// TIA Portal project "Lagerregal_3" (V20)

(* hardware
DEVICE "S7-1500/ET200MP-Station_1"  S7-1500 station
   slot 0: "Profilschiene_0"  Rack  6ES7 590-1***0-0AA0
   slot 1: "PLC_1"  CPU 1513-1 PN  6ES7 513-1AM03-0AB0  V4.0
      slot 3: "CPU-Display_1"  6ES7591-1AA00-0AA0
      slot 32768: "PROFINET-Schnittstelle_1"  X1
         slot 32769: "Port_1"  X1 P1
         slot 32770: "Port_2"  X1 P2
      slot 34817: "Virtual CP interface port_1"  Virtual CP interface port  Virtual CP interface port FW V4.0
   slot 2: "DI 16x24VDC BA_1"  DI 16x24VDC BA  6ES7 521-1BH10-0AA0  V1.1
   slot 3: "DQ 16x24VDC/0.5A ST_1"  DQ 16x24VDC/0.5A ST  6ES7 522-1BH00-0AB0  V2.0
   slot 4: "AI 8xU/I/R/RTD BA_2"  AI 8xU/I/R/RTD BA  6ES7 531-7QF00-0AB0  V1.0
   slot 5: "AI 8xU/I/R/RTD BA_1"  AI 8xU/I/R/RTD BA  6ES7 531-7QF00-0AB0  V1.0
DEVICE "HMI_1"  TP700 Comfort
   slot 0: "HMI_1"  TP700 Comfort  6AV2 124-0GC01-0AX0  17.0.0.0
   slot 1: "HMI_RT_1"  TP700 Comfort  6AV2 124-0GC01-0AX0  17.0.0.0
   slot 5: "HMI_1.IE_CP_1"  PROFINET Interface  17.0.0.0
      slot 1: "PROFINET Schnittstelle_1"  PROFINET Interface
         slot 1: "Port_1"  Port
         slot 2: "Port_2"  Port
   slot 7: "HMI_1.MPI/DP_CP_1"  MPI/DP Interface  17.0.0.0
*)

// ===== PLC "PLC_1"  CPU 1513-1 PN =====

VAR_GLOBAL   // PLC tag table "Standard-Variablentabelle"
   "Clock_Byte" AT %MB0 : Byte;
   "Clock_10Hz" AT %M0.0 : Bool;
   "Clock_5Hz" AT %M0.1 : Bool;
   "Clock_2.5Hz" AT %M0.2 : Bool;
   "Clock_2Hz" AT %M0.3 : Bool;
   "Clock_1.25Hz" AT %M0.4 : Bool;
   "Clock_1Hz" AT %M0.5 : Bool;
   "Clock_0.625Hz" AT %M0.6 : Bool;
   "Clock_0.5Hz" AT %M0.7 : Bool;
END_VAR

VAR_GLOBAL CONSTANT   // PLC tag table "Standard-Variablentabelle"
   "Fachhoehe" : Int := 4800;
   "Fachbreite" : Int := 2962;
   "Offset-Z" : Int := 1800;
   "Offset-X" : Int := 3952;
   "Faecher_pro_Zeile" : Int := 9;
   "Faecher_pro_Spalte" : Int := 6;
   "Anheben_Absenken" : Int := 1000;
END_VAR

VAR_GLOBAL   // PLC tag table "Eingaenge"
   "S1" AT %I0.0 : Bool;   // Not-Aus
   "S2" AT %I0.1 : Bool;   // Anlage ein
   "S3" AT %I0.2 : Bool;   // Starttaster
   "1B1" AT %I0.3 : Bool;   // Sensor 1. Einlassband Anfang
   "1B2" AT %I0.4 : Bool;   // Sensor 1. Einlassband Ende
   "2B1" AT %I0.5 : Bool;   // Sensor 2. Einlassband Anfang
   "2B2" AT %I0.6 : Bool;   // Sensor 2. Einlassband Ende
   "3B1" AT %I0.7 : Bool;   // Sensor 3. Einlassband
   "4B1" AT %I1.0 : Bool;   // Sensor 1. Auslassband
   "5B1" AT %I1.1 : Bool;   // Sensor 2. Auslassband
   "6B1" AT %I1.2 : Bool;   // Endlage Gabel-Kran 1 (links)
   "6B2" AT %I1.3 : Bool;   // Endlage Gabel-Kran 1 (rechts)
   "6B3" AT %I1.4 : Bool;   // Endlage Gabel-Kran 1 (mitte)
   "7B1" AT %I1.5 : Bool;   // Endlage Gabel-Kran 2 (links)
   "7B2" AT %I1.6 : Bool;   // Endlage Gabel-Kran 2 (rechts)
   "7B3" AT %I1.7 : Bool;   // Endlage Gabel-Kran 2 (mitte)
   "2B3" AT %EW30 : Int;   // Kamera am Einlass (Bauteilerkennung)
   "6B4" AT %EW32 : Int;   // X-Achse Kran 1 Ist-Pos
   "6B5" AT %EW34 : Int;   // Z-Achse Kran 1 Ist-Pos
   "7B4" AT %EW36 : Int;   // X-Achse Kran 2 Ist-Pos
   "7B5" AT %EW38 : Int;   // Z-Achse Kran 2 Ist-Pos
END_VAR

VAR_GLOBAL   // PLC tag table "Ausgaenge"
   "H3" AT %Q0.2 : Bool;   // Starttasterleuchte
   "1M1" AT %Q0.3 : Bool;   // 1. Einlassband
   "2M1" AT %Q0.5 : Bool;   // 2. Einlassband
   "3M1" AT %Q0.7 : Bool;   // 3. Einlassband
   "4M1" AT %Q1.0 : Bool;   // 1. Auslassband
   "5M1" AT %Q1.1 : Bool;   // 2. Auslassband
   "6M1" AT %Q1.2 : Bool;   // Gabel-Kran 1 (links)
   "6M2" AT %Q1.3 : Bool;   // Gabel-Kran 1 (rechts)
   "7M1" AT %Q1.5 : Bool;   // Gabel-Kran 2 (links)
   "7M2" AT %Q1.6 : Bool;   // Gabel-Kran 2 (rechts)
   "6M4" AT %AW32 : Int;   // X-Achse Kran 1 Soll-Pos
   "6M5" AT %AW34 : Int;   // Z-Achse Kran 1 Soll-Pos
   "7M4" AT %AW36 : Int;   // X-Achse Kran 2 Soll-Pos
   "7M5" AT %AW38 : Int;   // Z-Achse Kran 2 Soll-Pos
END_VAR

TYPE "typKran_Pos"
   STRUCT
      "X-Ist" : Int;
      "X-Soll" : Int;
      "Z-Ist" : Int;
      "Z-Soll" : Int;
   END_STRUCT;
END_TYPE

TYPE "typLagerplatz"
   STRUCT
      Flags : Struct
         Belegt : Bool;
         In_Benutzung : Bool;
      END_STRUCT;
   END_STRUCT;
END_TYPE

TYPE "typSchritte"
   STRUCT
      Schritt_Init : Bool;
      Kran : Struct
         Schritt_1 : Bool;
         Schritt_2 : Bool;
         Schritt_3 : Bool;
         Schritt_4 : Bool;
         Schritt_5 : Bool;
      END_STRUCT;
      Kran_Beladen : Struct
         Schritt_1 : Bool;
         Schritt_2 : Bool;
         Schritt_3 : Bool;
         Schritt_4 : Bool;
      END_STRUCT;
      Kran_Entladen : Struct
         Schritt_1 : Bool;
         Schritt_2 : Bool;
         Schritt_3 : Bool;
         Schritt_4 : Bool;
      END_STRUCT;
   END_STRUCT;
END_TYPE

DATA_BLOCK "IDB_Anlage"   // DB1
{ S7_Optimized_Access := 'TRUE' }
VERSION : 0.1
// stored: InstanceOfName Ein_Anlage
"Ein_Anlage"
BEGIN
END_DATA_BLOCK

DATA_BLOCK "IDB_Kran_beladen"   // DB2
{ S7_Optimized_Access := 'TRUE' }
VERSION : 0.1
// stored: InstanceOfName FC_Kran_beladen
"FC_Kran_beladen"
BEGIN
END_DATA_BLOCK

DATA_BLOCK "IDB_HMI"   // DB20
{ S7_Optimized_Access := 'TRUE' }
VERSION : 0.1
// stored: InstanceOfName Ein_HMI
"Ein_HMI"
BEGIN
END_DATA_BLOCK

DATA_BLOCK "IDB_Einrichtbetrieb"   // DB30
{ S7_Optimized_Access := 'TRUE' }
VERSION : 0.1
// stored: InstanceOfName Prog_Einrichtbetrieb
"Prog_Einrichtbetrieb"
BEGIN
END_DATA_BLOCK

DATA_BLOCK "IDB_Automatik_einlagern"   // DB50
{ S7_Optimized_Access := 'TRUE' }
VERSION : 0.1
// stored: InstanceOfName Prog_Automatik_einlagern
"Prog_Automatik_einlagern"
BEGIN
END_DATA_BLOCK

DATA_BLOCK "HMI_Schnittstelle"   // DB100
{ S7_Optimized_Access := 'TRUE' }
VERSION : 0.1
   VAR
      Betriebsart : Struct
         Hand : Bool;
         Automatik : Bool;
         Einrichten : Bool;
         Grundstellung_Einlagern : Bool;
         Grundstellung_Auslagern : Bool;
         Regalplatz_frei : Bool;
      END_STRUCT;
      Automatik_EIN : Struct
         Calc_POS_X : Int;
         Calc_POS_Z : Int;
         Schrittnummer : Int;
         FachNr : Int := 1;
      END_STRUCT;
      Schrittnummer : UDInt;
      Fach : Int;
      Fach_ansteuern : Bool;
      Eingaenge : Struct
         S1 : Bool;
         S2 : Bool;
         S3 : Bool;
         "1B1" : Bool;
         "1B2" : Bool;
         "2B1" : Bool;
         "2B2" : Bool;
         "3B1" : Bool;
         "4B1" : Bool;
         "5B1" : Bool;
         "6B1" : Bool;
         "6B2" : Bool;
         "6B3" : Bool;
         "7B1" : Bool;
         "7B2" : Bool;
         "7B3" : Bool;
      END_STRUCT;
      Ausgaenge : Struct
         H1 : Bool;
         "1M1" : Bool;
         "2M1" : Bool;
         "3M1" : Bool;
         "4M1" : Bool;
         "5M1" : Bool;
         "6M1" : Bool;
         "6M2" : Bool;
         "7M1" : Bool;
         "7M2" : Bool;
      END_STRUCT;
      Kraene : Struct
         Kran_1 : Struct
            Kran_Pos : "typKran_Pos";
            Gabel : Struct
               Links : Bool;
               Rechts : Bool;
            END_STRUCT;
            Schritt_Kran : Int;
            Schritt_Beladen : Int;
            Schritt_Entladen : Int;
            Home : Bool;
            Steht : Bool;
            Beladen : Bool;
         END_STRUCT;
         Kran_2 : Struct
            Kran_Pos : "typKran_Pos";
            Gabel : Struct
               Links : Bool;
               Rechts : Bool;
            END_STRUCT;
            Schritt_Kran : Int;
            Schritt_Beladen : Int;
            Schritt_Entladen : Int;
            Home : Bool;
            Steht : Bool;
            Beladen : Bool;
         END_STRUCT;
      END_STRUCT;
      HMI : Struct
         "X-Pos" : Bool;
         "X-Neg" : Bool;
         "Z-Pos" : Bool;
         "Z-Neg" : Bool;
         Inkrement : UInt;
      END_STRUCT;
   END_VAR
BEGIN
END_DATA_BLOCK

DATA_BLOCK "Warenlager"   // DB101
{ S7_Optimized_Access := 'TRUE' }
VERSION : 0.1
   VAR
      Lager : Array[1..54] of "typLagerplatz";
   END_VAR
BEGIN
END_DATA_BLOCK

FUNCTION_BLOCK "Ein_Anlage"   // FB1, FBD
{ S7_Optimized_Access := 'TRUE' }
VERSION : 0.1
   VAR
      NTRIG_MDB_1B2 : F_TRIG;
      NTRIG_MDB_2B2 : F_TRIG;
      NTRIG_MDB_5B1 : F_TRIG;
   END_VAR
BEGIN

REGION Network 1: Schalter einlesen
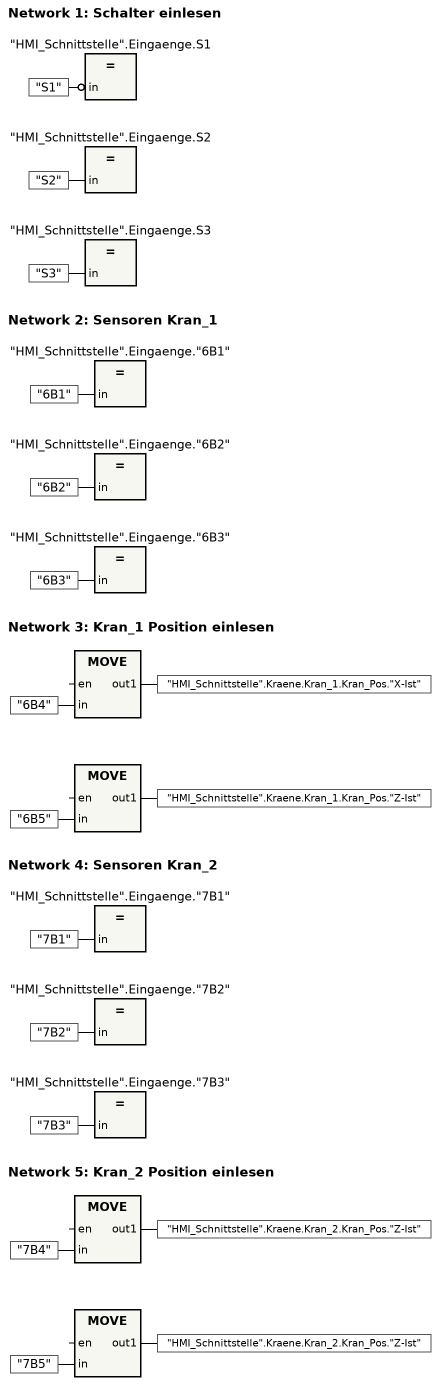
   "HMI_Schnittstelle".Eingaenge.S1 := NOT "S1";
   "HMI_Schnittstelle".Eingaenge.S2 := "S2";
   "HMI_Schnittstelle".Eingaenge.S3 := "S3";
END_REGION

REGION Network 2: Sensoren Kran_1
   "HMI_Schnittstelle".Eingaenge."6B1" := "6B1";
   "HMI_Schnittstelle".Eingaenge."6B2" := "6B2";
   "HMI_Schnittstelle".Eingaenge."6B3" := "6B3";
END_REGION

REGION Network 3: Kran_1 Position einlesen
   "HMI_Schnittstelle".Kraene.Kran_1.Kran_Pos."X-Ist" := "6B4";
   "HMI_Schnittstelle".Kraene.Kran_1.Kran_Pos."Z-Ist" := "6B5";
END_REGION

REGION Network 4: Sensoren Kran_2
   "HMI_Schnittstelle".Eingaenge."7B1" := "7B1";
   "HMI_Schnittstelle".Eingaenge."7B2" := "7B2";
   "HMI_Schnittstelle".Eingaenge."7B3" := "7B3";
END_REGION

REGION Network 5: Kran_2 Position einlesen
   "HMI_Schnittstelle".Kraene.Kran_2.Kran_Pos."Z-Ist" := "7B4";
   "HMI_Schnittstelle".Kraene.Kran_2.Kran_Pos."Z-Ist" := "7B5";
END_REGION

REGION Network 6: Sensoren Einlass
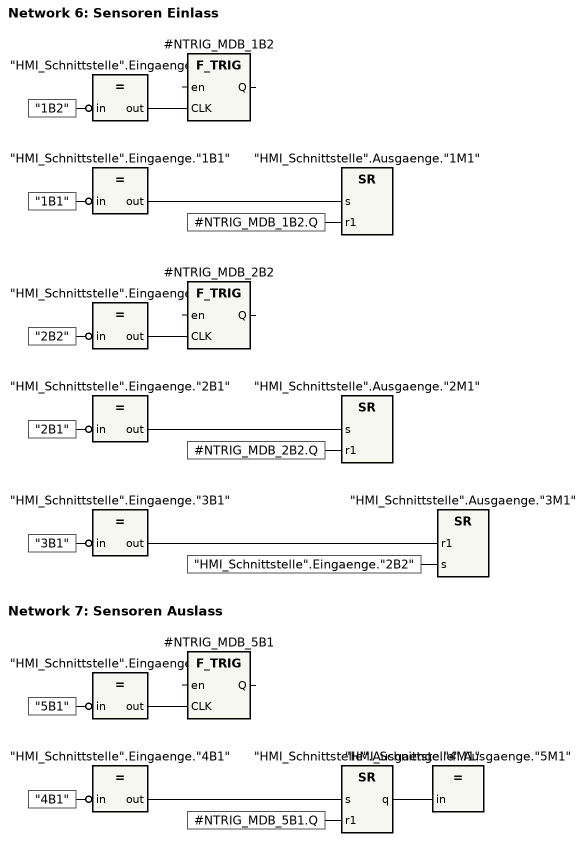
   "HMI_Schnittstelle".Eingaenge."1B2" := NOT "1B2";
   #NTRIG_MDB_1B2(CLK := NOT "1B2");   // F_TRIG
   "HMI_Schnittstelle".Eingaenge."1B1" := NOT "1B1";
   IF NOT "1B1" THEN
       "HMI_Schnittstelle".Ausgaenge."1M1" := TRUE;   // SR flip-flop
   END_IF;
   IF #NTRIG_MDB_1B2.Q THEN "HMI_Schnittstelle".Ausgaenge."1M1" := FALSE; END_IF;
   "HMI_Schnittstelle".Eingaenge."2B2" := NOT "2B2";
   #NTRIG_MDB_2B2(CLK := NOT "2B2");   // F_TRIG
   "HMI_Schnittstelle".Eingaenge."2B1" := NOT "2B1";
   IF NOT "2B1" THEN
       "HMI_Schnittstelle".Ausgaenge."2M1" := TRUE;   // SR flip-flop
   END_IF;
   IF #NTRIG_MDB_2B2.Q THEN "HMI_Schnittstelle".Ausgaenge."2M1" := FALSE; END_IF;
   "HMI_Schnittstelle".Eingaenge."3B1" := NOT "3B1";
   IF "HMI_Schnittstelle".Eingaenge."2B2" THEN
       "HMI_Schnittstelle".Ausgaenge."3M1" := TRUE;   // SR flip-flop
   END_IF;
   IF NOT "3B1" THEN "HMI_Schnittstelle".Ausgaenge."3M1" := FALSE; END_IF;
END_REGION

REGION Network 7: Sensoren Auslass
   "HMI_Schnittstelle".Eingaenge."5B1" := NOT "5B1";
   #NTRIG_MDB_5B1(CLK := NOT "5B1");   // F_TRIG
   "HMI_Schnittstelle".Eingaenge."4B1" := NOT "4B1";
   IF NOT "4B1" THEN
       "HMI_Schnittstelle".Ausgaenge."4M1" := TRUE;   // SR flip-flop
   END_IF;
   IF #NTRIG_MDB_5B1.Q THEN "HMI_Schnittstelle".Ausgaenge."4M1" := FALSE; END_IF;
   "HMI_Schnittstelle".Ausgaenge."5M1" := "HMI_Schnittstelle".Ausgaenge."4M1";
END_REGION
END_FUNCTION_BLOCK

FUNCTION_BLOCK "FC_Kran_beladen"   // FB2, FBD
{ S7_Optimized_Access := 'TRUE' }
VERSION : 0.1
   VAR_INPUT
      "eKran_Z-Ist" : Int;
      eSchrittnummer : Int;
   END_VAR
   VAR_OUTPUT
      aGabel : Bool;
      aBeladen : Bool;
      "aKran_Z-Soll" : Int;
   END_VAR
   VAR
      PTRIG_Schritt2 : Bool;
   END_VAR
   VAR_TEMP   // added for the SCL form of the ladder/FBD networks
      _w1 : Bool;
      _w2 : Bool;
   END_VAR
BEGIN

REGION Network 1: Gabel zur Seite ausfahren
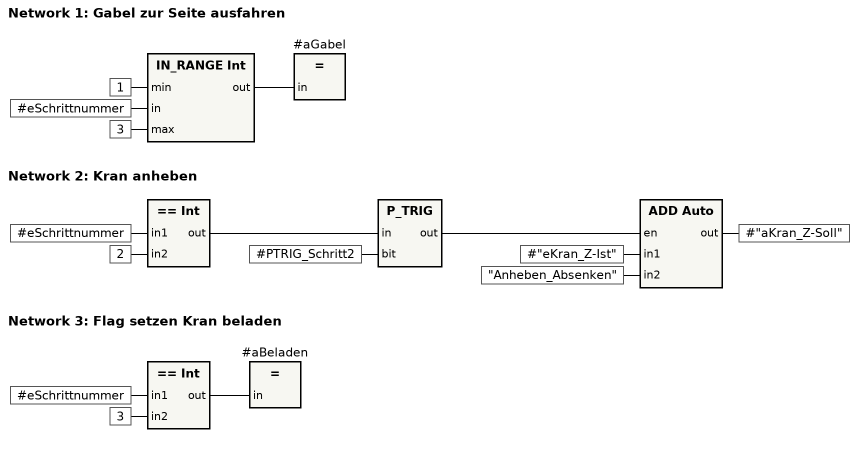
   #aGabel := (1 <= #eSchrittnummer) AND (#eSchrittnummer <= 3);
END_REGION

REGION Network 2: Kran anheben
   #_w1 := #eSchrittnummer = 2;
   #_w2 := #_w1 AND NOT #PTRIG_Schritt2;   // rising edge
   #PTRIG_Schritt2 := #_w1;
   IF #_w2 THEN #"aKran_Z-Soll" := #"eKran_Z-Ist" + "Anheben_Absenken"; END_IF;
END_REGION

REGION Network 3: Flag setzen Kran beladen
   #aBeladen := #eSchrittnummer = 3;
END_REGION
END_FUNCTION_BLOCK

FUNCTION_BLOCK "FC_Kran_entladen"   // FB3, FBD
{ S7_Optimized_Access := 'TRUE' }
VERSION : 0.1
   VAR_INPUT
      "eKran_Z-Ist" : Int;
      eSchrittnummer : Int;
   END_VAR
   VAR_OUTPUT
      aGabel : Bool;
      aBeladen : Bool;
      "aKran_Z-Soll" : Int;
   END_VAR
   VAR
      PTRIG_Schritt2 : Bool;
   END_VAR
   VAR_TEMP   // added for the SCL form of the ladder/FBD networks
      _w1 : Bool;
      _w2 : Bool;
   END_VAR
BEGIN

REGION Network 1: Gabel zur Seite ausfahren
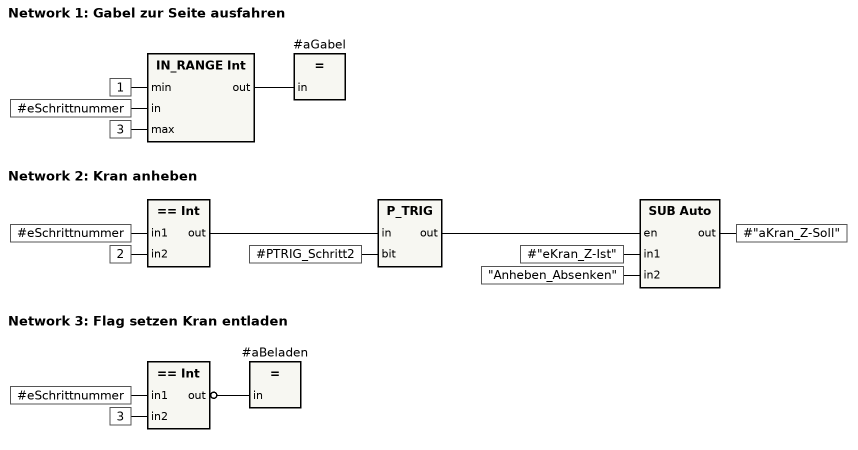
   #aGabel := (1 <= #eSchrittnummer) AND (#eSchrittnummer <= 3);
END_REGION

REGION Network 2: Kran anheben
   #_w1 := #eSchrittnummer = 2;
   #_w2 := #_w1 AND NOT #PTRIG_Schritt2;   // rising edge
   #PTRIG_Schritt2 := #_w1;
   IF #_w2 THEN #"aKran_Z-Soll" := #"eKran_Z-Ist" - "Anheben_Absenken"; END_IF;
END_REGION

REGION Network 3: Flag setzen Kran entladen
   #aBeladen := NOT (#eSchrittnummer = 3);
END_REGION
END_FUNCTION_BLOCK

FUNCTION_BLOCK "Ein_HMI"   // FB20, FBD
{ S7_Optimized_Access := 'TRUE' }
VERSION : 0.1
BEGIN
END_FUNCTION_BLOCK

FUNCTION_BLOCK "Bandsteuerung"   // FB21, FBD
{ S7_Optimized_Access := 'TRUE' }
VERSION : 0.1
   VAR
      RTRIG_Palette_geladen : R_TRIG;
      FTRIG_Palette_an_Band1_Ende : F_TRIG;
      Band_belegt : Bool;
   END_VAR
BEGIN

REGION Network 1 (SCL): Flankenabfragen
   #RTRIG_Palette_geladen(CLK:="HMI_Schnittstelle".Automatik_EIN.Schrittnummer = 5);
   #FTRIG_Palette_an_Band1_Ende(CLK:="HMI_Schnittstelle".Eingaenge."1B2");
END_REGION

REGION Network 2: Band belegt
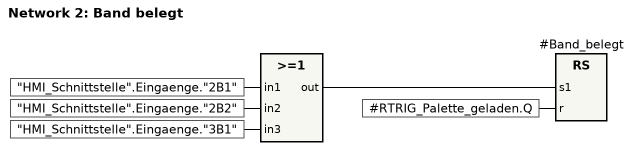
   IF #RTRIG_Palette_geladen.Q THEN
       #Band_belegt := FALSE;   // RS flip-flop
   END_IF;
   IF "HMI_Schnittstelle".Eingaenge."2B1" OR "HMI_Schnittstelle".Eingaenge."2B2" OR "HMI_Schnittstelle".Eingaenge."3B1" THEN
       #Band_belegt := TRUE;
   END_IF;
END_REGION
END_FUNCTION_BLOCK

FUNCTION_BLOCK "Prog_Einrichtbetrieb"   // FB30, FBD
{ S7_Optimized_Access := 'TRUE' }
VERSION : 0.1
   VAR
      "PTRIG_MDB_X-Pos" : R_TRIG;
      "PTRIG_MDB_X-Neg" : R_TRIG;
      "PTRIG_MDB_Z-Pos" : R_TRIG;
      "PTRIG_MDB_Z-Neg" : R_TRIG;
   END_VAR
BEGIN

REGION Network 1: Button Flanken erfassen
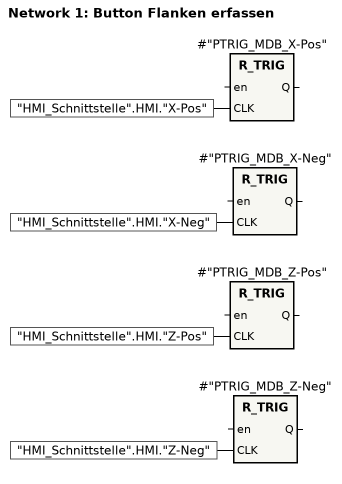
   #"PTRIG_MDB_X-Pos"(CLK := "HMI_Schnittstelle".HMI."X-Pos");   // R_TRIG
   #"PTRIG_MDB_X-Neg"(CLK := "HMI_Schnittstelle".HMI."X-Neg");   // R_TRIG
   #"PTRIG_MDB_Z-Pos"(CLK := "HMI_Schnittstelle".HMI."Z-Pos");   // R_TRIG
   #"PTRIG_MDB_Z-Neg"(CLK := "HMI_Schnittstelle".HMI."Z-Neg");   // R_TRIG
END_REGION

REGION Network 2 (SCL): Achsen inkrementieren
   // X-Achse Inkrementieren
   IF #"PTRIG_MDB_X-Pos".Q THEN
       "HMI_Schnittstelle".Kraene.Kran_1.Kran_Pos."X-Soll" += UINT_TO_INT("HMI_Schnittstelle".HMI.Inkrement);
   END_IF;

   IF #"PTRIG_MDB_X-Neg".Q THEN
       "HMI_Schnittstelle".Kraene.Kran_1.Kran_Pos."X-Soll" -= UINT_TO_INT("HMI_Schnittstelle".HMI.Inkrement);
   END_IF;


   // Z-Achse Inkrementieren
   IF #"PTRIG_MDB_Z-Pos".Q THEN
       "HMI_Schnittstelle".Kraene.Kran_1.Kran_Pos."Z-Soll" += UINT_TO_INT("HMI_Schnittstelle".HMI.Inkrement);
   END_IF;

   IF #"PTRIG_MDB_Z-Neg".Q THEN
       "HMI_Schnittstelle".Kraene.Kran_1.Kran_Pos."Z-Soll" -= UINT_TO_INT("HMI_Schnittstelle".HMI.Inkrement);
   END_IF;
END_REGION
END_FUNCTION_BLOCK

FUNCTION_BLOCK "Prog_Automatik_einlagern"   // FB50, FBD
{ S7_Optimized_Access := 'TRUE' }
VERSION : 0.1
   VAR
      MDB_Schrittkette_einlagern : "Prog_Schrittkette";
      FTRIG_Palette_eingelagert : F_TRIG;
   END_VAR
   VAR_TEMP
      tmpPalette_abgelegt : Int;
   END_VAR
BEGIN

REGION Network 1: Lagerplatz frei
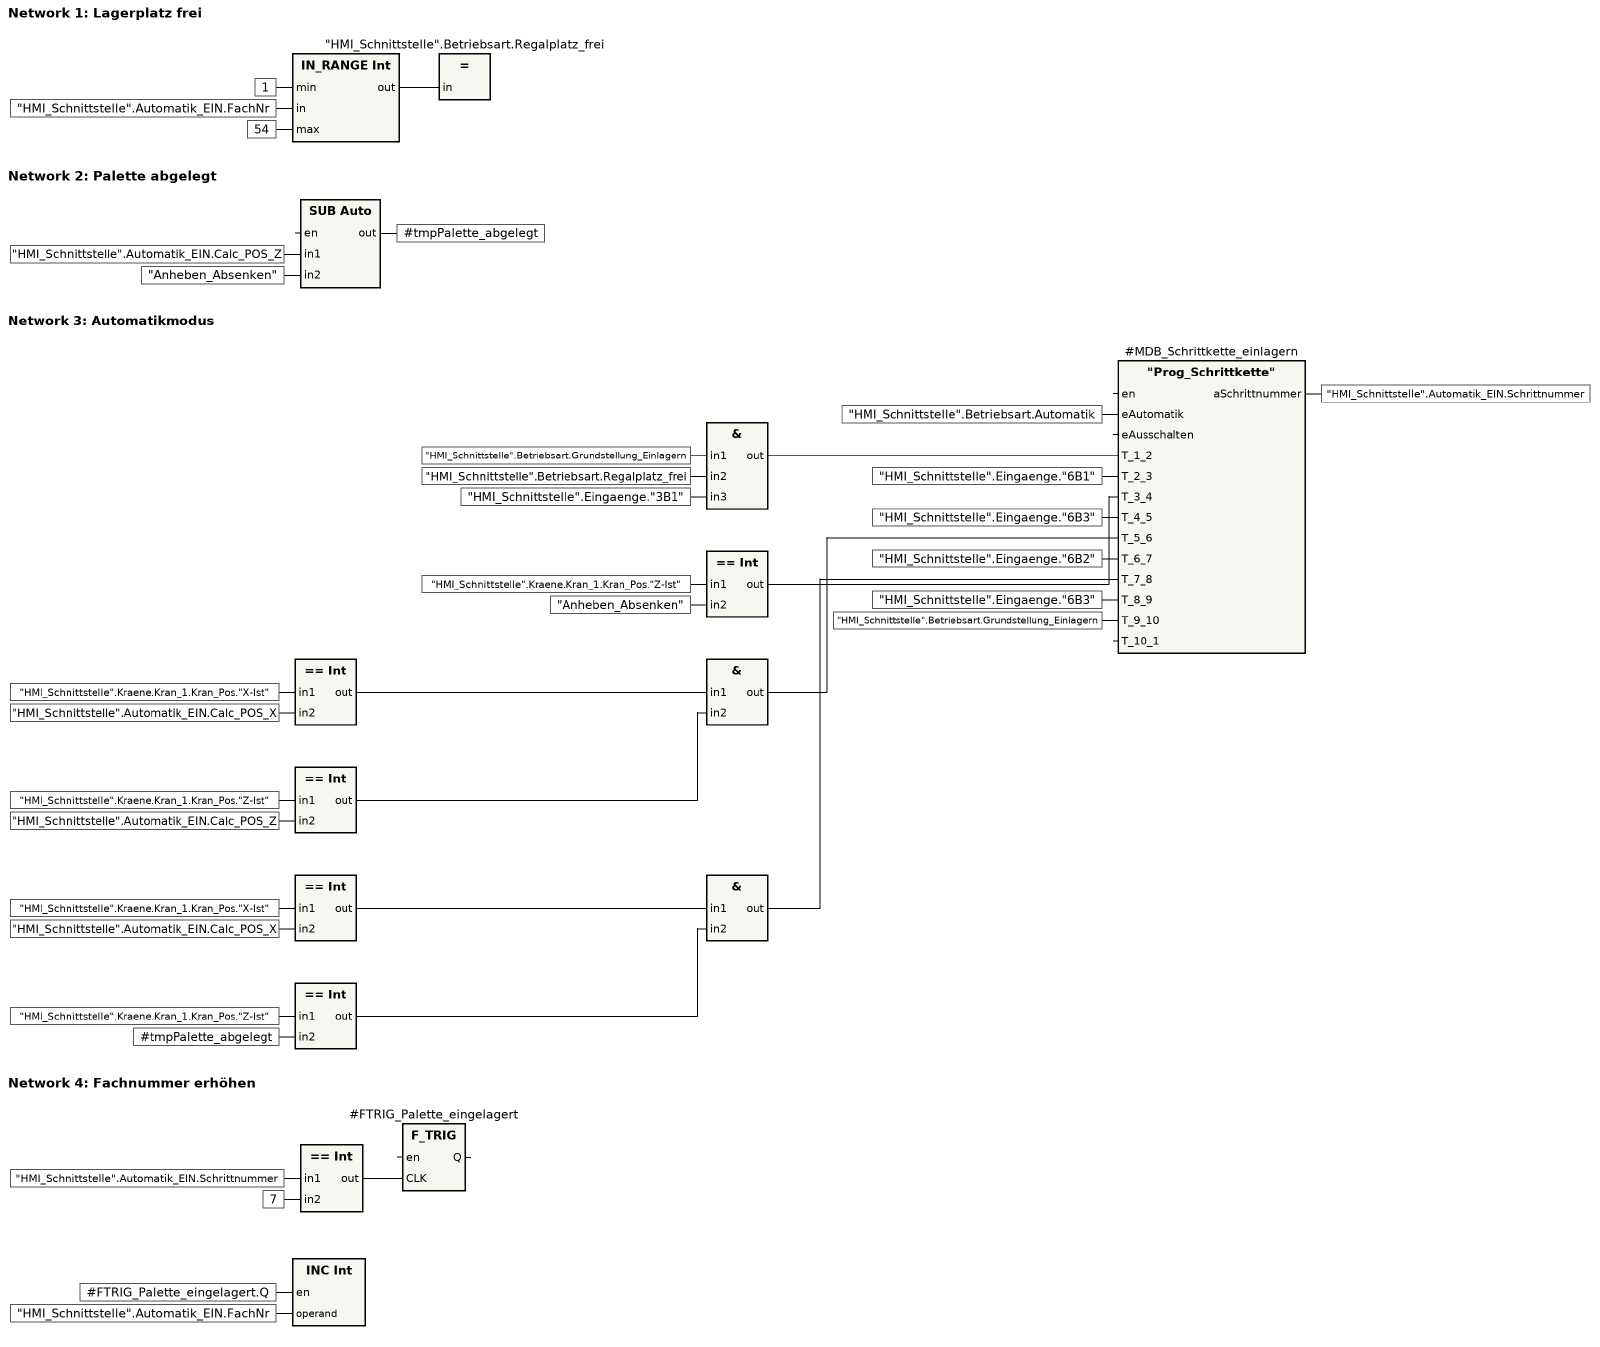
   "HMI_Schnittstelle".Betriebsart.Regalplatz_frei := (1 <= "HMI_Schnittstelle".Automatik_EIN.FachNr) AND ("HMI_Schnittstelle".Automatik_EIN.FachNr <= 54);
END_REGION

REGION Network 2: Palette abgelegt
   #tmpPalette_abgelegt := "HMI_Schnittstelle".Automatik_EIN.Calc_POS_Z - "Anheben_Absenken";
END_REGION

REGION Network 3: Automatikmodus
   #MDB_Schrittkette_einlagern(eAutomatik := "HMI_Schnittstelle".Betriebsart.Automatik,   // "Prog_Schrittkette"
                           T_1_2 := "HMI_Schnittstelle".Betriebsart.Grundstellung_Einlagern AND "HMI_Schnittstelle".Betriebsart.Regalplatz_frei AND "HMI_Schnittstelle".Eingaenge."3B1",
                           T_2_3 := "HMI_Schnittstelle".Eingaenge."6B1",
                           T_3_4 := "HMI_Schnittstelle".Kraene.Kran_1.Kran_Pos."Z-Ist" = "Anheben_Absenken",
                           T_4_5 := "HMI_Schnittstelle".Eingaenge."6B3",
                           T_5_6 := ("HMI_Schnittstelle".Kraene.Kran_1.Kran_Pos."X-Ist" = "HMI_Schnittstelle".Automatik_EIN.Calc_POS_X) AND ("HMI_Schnittstelle".Kraene.Kran_1.Kran_Pos."Z-Ist" = "HMI_Schnittstelle".Automatik_EIN.Calc_POS_Z),
                           T_6_7 := "HMI_Schnittstelle".Eingaenge."6B2",
                           T_7_8 := ("HMI_Schnittstelle".Kraene.Kran_1.Kran_Pos."X-Ist" = "HMI_Schnittstelle".Automatik_EIN.Calc_POS_X) AND ("HMI_Schnittstelle".Kraene.Kran_1.Kran_Pos."Z-Ist" = #tmpPalette_abgelegt),
                           T_8_9 := "HMI_Schnittstelle".Eingaenge."6B3",
                           T_9_10 := "HMI_Schnittstelle".Betriebsart.Grundstellung_Einlagern,
                           aSchrittnummer => "HMI_Schnittstelle".Automatik_EIN.Schrittnummer);
END_REGION

REGION Network 4: Fachnummer erhöhen
   #FTRIG_Palette_eingelagert(CLK := "HMI_Schnittstelle".Automatik_EIN.Schrittnummer = 7);   // F_TRIG
   IF #FTRIG_Palette_eingelagert.Q THEN
       "HMI_Schnittstelle".Automatik_EIN.FachNr := "HMI_Schnittstelle".Automatik_EIN.FachNr + 1;
   END_IF;
END_REGION
END_FUNCTION_BLOCK

FUNCTION_BLOCK "Prog_Schrittkette"   // FB1234, FBD
{ S7_Optimized_Access := 'TRUE' }